HMI tags "BC_HMI_Tags"
   "10 DI_DATA_E131_OK" : Bool = PLC "20_TANKS_IP_DATA".RIO_03.FIRST_TANK.USD_FLOW AT %DB1.DBX0.0, 1 s
   "10 DI_DATA_E131_SHTDN" : Bool = PLC "10 DI_DATA".E131_SHTDN AT %DB1.DBX0.0, 1 s
   "103_Main_Burner_DB_DN_OK(1)" : Bool = PLC "103_Main_Burner_DB".DN_OK AT %DB1.DBX0.0, 1 s
   "10 DI_DATA_FD001_OK" : Bool = PLC "10 DI_DATA".FD001_OK AT %DB1.DBX0.0, 1 s
   "10 DI_DATA_FD001_PWR_OK" : Bool = PLC "10 DI_DATA".FD001_PWR_OK AT %DB1.DBX0.0, 1 s
   "10 DI_DATA_FS115(1)" : Bool = PLC "10 DI_DATA".FS115 AT %DB1.DBW0, 1 s
   "10 DI_DATA_FS123" : Bool = PLC "10 DI_DATA".FS123 AT %DB1.DBX0.0, 1 s
   "10 DI_DATA_FS317" : Bool = PLC "10 DI_DATA".FS317 AT %DB1.DBX0.0, 1 s
   "10 DI_DATA_FS320" : Bool = PLC "10 DI_DATA".FS320 AT %DB1.DBX0.0, 1 s
   "10 DI_DATA_ESD_OK" : Bool = PLC "10 DI_DATA".ESD_OK AT %DB1.DBX0.0, 1 s
   "10 DI_DATA_P301_ENBLD" : Bool = PLC "10 DI_DATA".P301_ENBLD AT %DB1.DBX0.0, 1 s
   "10 DI_DATA_R2_SPR_DI_1_6" : Bool = PLC "10 DI_DATA".R2_SPR_DI_1_6 AT %DB1.DBX0.0, 1 s
   "10 DI_DATA_P301_TRIPPED(1)" : Bool = PLC "10 DI_DATA".P301_TRIPPED AT %DB1.DBX0.0, 1 s
   "10 DI_DATA_P305_ENBLD" : Bool = PLC "10 DI_DATA".P305_ENBLD AT %DB1.DBX0.0, 1 s
   "10 DI_DATA_P305_TRIPPED(1)" : Bool = PLC "10 DI_DATA".P305_TRIPPED AT %DB1.DBX0.0, 1 s
   "10 DI_DATA_PS101" : Bool = PLC "10 DI_DATA".PS101 AT %DB1.DBX0.0, 1 s
   "10 DI_DATA_R2_SPR_DI_0_2" : Bool = PLC "10 DI_DATA".R2_SPR_DI_0_2 AT %DB1.DBX0.0, 1 s
   "10 DI_DATA_R2_SPR_DI_0_3" : Bool = PLC "10 DI_DATA".R2_SPR_DI_0_3 AT %DB1.DBX0.0, 1 s
   "10 DI_DATA_TS403_FAULT" : Bool = PLC "10 DI_DATA".TS403_FAULT AT %DB1.DBX0.0, 1 s
   "10 DI_DATA_X001_PWR_OK" : Bool = PLC "10 DI_DATA".X001_PWR_OK AT %DB1.DBX0.0, 1 s
   "102_Pilot_Burner_DB_FLM_DET" : Bool = PLC "102_Pilot_Burner_DB".FLM_DET AT %DB1.DBX0.0, 100 ms
   "104_Pilot_Purge_DB_DN_OK" : Bool = PLC "104_Pilot_Purge_DB".DN_OK AT %DB1.DBX0.0, 1 s
   "10 DI_DATA_E600_NOK" : Bool = PLC "10 DI_DATA".E600_NOK AT %DB1.DBX0.0, 1 s
   "10 DI_DATA_E600_HIHI" : Bool = PLC "10 DI_DATA".E600_HIHI AT %DB1.DBX0.0, 1 s
   "10 DI_DATA_E600_LOLO" : Bool = PLC "10 DI_DATA".E600_LOLO AT %DB1.DBX0.0, 1 s
   "10 DI_DATA_E600_PWR_OK" : Bool = PLC "10 DI_DATA".E600_PWR_OK AT %DB1.DBX0.0, 1 s
   "10 DI_DATA_E700_PWR_OK" : Bool = PLC "10 DI_DATA".E700_PWR_OK AT %DB1.DBX0.0, 1 s
   "10 DI_DATA_E700_OPACITY" : Bool = PLC "10 DI_DATA".E700_OPACITY AT %DB1.DBX0.0, 1 s
   "10 DI_DATA_TS403_FAULT(1)" : Bool = PLC "10 DI_DATA".TS403_FAULT AT %DB1.DBX0.0, 1 s
   "10 DI_DATA_TS006" : Bool = PLC "10 DI_DATA".TS006 AT %DB1.DBX0.0, 1 s
   "10 DI_DATA_S2_8K1_OK" : Bool = PLC "10 DI_DATA".S2_8K1_OK AT %DB1.DBX0.0, 1 s
   "10 DI_DATA_E131_WRNG" : Bool = PLC "10 DI_DATA".E131_WRNG AT %DB1.DBX0.0, 1 s
   "10 DI_DATA_R2_SPR_DI_3_2" : Bool = PLC "10 DI_DATA".R2_SPR_DI_3_2 AT %DB1.DBX0.0, 1 s
   "10 DI_DATA_R2_SPR_DI_3_7" : Bool = PLC "10 DI_DATA".R2_SPR_DI_3_7 AT %DB1.DBX0.0, 1 s
   "10 DI_DATA_LS001" : Bool = PLC "10 DI_DATA".LS001 AT %DB1.DBX0.0, 1 s
   "10 DI_DATA_P305_TRIPPED" : Bool = PLC "10 DI_DATA".P305_TRIPPED AT %DB1.DBX0.0, 1 s
   "10 DI_DATA_P305_ENBLD(1)" : Bool = PLC "10 DI_DATA".P305_ENBLD AT %DB1.DBX0.0, 1 s
   "84_Setpoints_PIT113_High" : Real = PLC "84_Setpoints".PIT113_High AT %DB1.DBD0, 1 s
   "84_Setpoints_PIT113_HighHigh" : Real = PLC "84_Setpoints".PIT113_HighHigh AT %DB1.DBD0, 1 s
   "84_Setpoints_PIT113_Pilot_Target" : Real = PLC "84_Setpoints".PIT113_Pilot_Target AT %DB1.DBX0.0, 1 s
   "84_Setpoints_PIT204_High(2)" : Real = PLC "84_Setpoints".PIT204_High, 1 s
   "84_Setpoints_PIT204_HighHigh(2)" : Real = PLC "84_Setpoints".PIT204_HighHigh, 1 s
   "84_Setpoints_PIT204_Low(2)" : Real = PLC "84_Setpoints".PIT204_Low, 1 s
   "84_Setpoints_PIT204_LowLow(2)" : Real = PLC "84_Setpoints".PIT204_LowLow, 1 s
   "84_Setpoints_PIT205_High" : Real = PLC "2084_Setpoints"."TX427 Star DO Lo" AT %DB1.DBD0, 1 s
   "84_Setpoints_PIT205_HighHigh" : Real = PLC "84_Setpoints".PIT205_HighHigh AT %DB1.DBD0, 1 s
   "84_Setpoints_PIT205_Low" : Real = PLC "84_Setpoints".PIT205_Low AT %DB1.DBD0, 1 s
   "84_Setpoints_PIT205_LowLow" : Real = PLC "84_Setpoints".PIT205_LowLow AT %DB1.DBD0, 1 s
   "84_Setpoints_PIT205_Target" : Real = PLC "84_Setpoints".PIT205_Target AT %DB1.DBX0.0, 1 s
   "84_Setpoints_PIT113_Low" : Real = PLC "84_Setpoints".PIT113_Low AT %DB1.DBD0, 1 s
   "84_Setpoints_PIT113_LowLow" : Real = PLC "84_Setpoints".PIT113_LowLow AT %DB1.DBD0, 1 s
   "84_Setpoints_TIT202_High" : Real = PLC "84_Setpoints".TIT202_High AT %DB1.DBD0, 1 s
   "84_Setpoints_TIT202_HighHigh" : Real = PLC "84_Setpoints".TIT202_HighHigh AT %DB1.DBD0, 1 s
   "84_Setpoints_TIT202_LowLow" : Real = PLC "84_Setpoints".TIT202_LowLow AT %DB1.DBD0, 1 s
   "84_Setpoints_TIT202_Low" : Real = PLC "84_Setpoints".TIT202_Low AT %DB1.DBD0, 1 s
   "84_Setpoints_TX700_High" : Real = PLC "84_Setpoints".TX700_High AT %DB1.DBD0, 1 s
   "84_Setpoints_TX700_Low" : Real = PLC "84_Setpoints".TX700_Low AT %DB1.DBD0, 1 s
   "84_Setpoints_FD001_LowLow" : Real = PLC "84_Setpoints".FD001_LowLow AT %DB1.DBD0, 1 s
   "84_Setpoints_E600_BWT_High" : Real = PLC "84_Setpoints".E600_BWT_High AT %DB1.DBD0, 1 s
   "84_Setpoints_E600_BWT_Low" : Real = PLC "84_Setpoints".E600_BWT_Low AT %DB1.DBD0, 1 s
   "84_Setpoints_FD001_Low" : Real = PLC "84_Setpoints".FD001_Low AT %DB1.DBD0, 1 s
   "84_Setpoints_AT_O2_1_LowLow" : Real = PLC "84_Setpoints".AT_O2_1_LowLow AT %DB1.DBD0, 1 s
   "84_Setpoints_AT_O2_2_LowLow" : Real = PLC "84_Setpoints".AT_O2_2_LowLow AT %DB1.DBD0, 1 s
   "84_Setpoints_AT_O2_2_Low" : Real = PLC "84_Setpoints".AT_O2_2_Low AT %DB1.DBD0, 1 s
   "80_From_HMI_MAN_DQ_1_7(1)" : Bool = PLC "80_From_HMI".MAN_DQ_1_7 AT %DB1.DBX0.0, 1 s
   "80_From_HMI_MAN_DQ_1_6" : Bool = PLC "80_From_HMI".MAN_DQ_1_6 AT %DB1.DBX0.0, 1 s
   "80_From_HMI_MAN_DQ_1_5(1)" : Bool = PLC "80_From_HMI".MAN_DQ_1_5 AT %DB1.DBX0.0, 1 s
   "80_From_HMI_MAN_DQ_1_4(1)" : Bool = PLC "80_From_HMI".MAN_DQ_1_4 AT %DB1.DBX0.0, 1 s
   "80_From_HMI_MAN_DQ_1_3(1)" : Bool = PLC "80_From_HMI".MAN_DQ_1_3 AT %DB1.DBX0.0, 1 s
   "80_From_HMI_MAN_DQ_1_2(1)" : Bool = PLC "80_From_HMI".MAN_DQ_1_2 AT %DB1.DBX0.0, 1 s
   "80_From_HMI_MAN_DQ_1_1(1)" : Bool = PLC "80_From_HMI".MAN_DQ_1_1 AT %DB1.DBX0.0, 1 s
   "80_From_HMI_MAN_DQ_1_0" : Bool = PLC "80_From_HMI".MAN_DQ_1_0 AT %DB1.DBX0.0, 1 s
   "80_From_HMI_MAN_DQ_0_7" : Bool = PLC "80_From_HMI".MAN_DQ_0_7 AT %DB1.DBX0.0, 1 s
   "80_From_HMI_MAN_DQ_0_6(1)" : Bool = PLC "80_From_HMI".MAN_DQ_0_6 AT %DB1.DBX0.0, 1 s
   "80_From_HMI_MAN_DQ_0_5(1)" : Bool = PLC "80_From_HMI".MAN_DQ_0_5 AT %DB1.DBX0.0, 1 s
   "80_From_HMI_MAN_DQ_0_4(1)" : Bool = PLC "80_From_HMI".MAN_DQ_0_4 AT %DB1.DBX0.0, 1 s
   "80_From_HMI_MAN_DQ_0_3(1)" : Bool = PLC "80_From_HMI".MAN_DQ_0_3 AT %DB1.DBX0.0, 1 s
   "80_From_HMI_MAN_DQ_0_2(1)" : Bool = PLC "80_From_HMI".MAN_DQ_0_2 AT %DB1.DBX0.0, 1 s
   "80_From_HMI_MAN_DQ_0_1(1)" : Bool = PLC "80_From_HMI".MAN_DQ_0_1 AT %DB1.DBX0.0, 1 s
   "80_From_HMI_MAN_DQ_0_0(1)" : Bool = PLC "80_From_HMI".MAN_DQ_0_0 AT %DB1.DBX0.0, 1 s
   "16_AQ_Data_CV111_CNTRL" : Real = PLC "16_AQ_Data".CV111_CNTRL AT %DB1.DBD0, 1 s
   "14_DQ_Data_X001ControlOut" : Bool = PLC "14_DQ_Data".X001ControlOut AT %DB1.DBX0.0, 1 s
   "14_DQ_Data_R2_SPR_DQ_1_6" : Bool = PLC "14_DQ_Data".R2_SPR_DQ_1_6 AT %DB1.DBX0.0, 1 s
   "14_DQ_Data_R2_SPR_DQ_1_4" : Bool = PLC "14_DQ_Data".R2_SPR_DQ_1_4 AT %DB1.DBX0.0, 1 s
   "14_DQ_Data_R2_SPR_DQ_1_5" : Bool = PLC "14_DQ_Data".R2_SPR_DQ_1_5 AT %DB1.DBX0.0, 1 s
   "14_DQ_Data_R2_SPR_DQ_1_3" : Bool = PLC "14_DQ_Data".R2_SPR_DQ_1_3 AT %DB1.DBX0.0, 1 s
   "14_DQ_Data_R2_SPR_DQ_1_2" : Bool = PLC "14_DQ_Data".R2_SPR_DQ_1_2 AT %DB1.DBX0.0, 1 s
   "14_DQ_Data_P305ControlOut" : Bool = PLC "14_DQ_Data".P305ControlOut AT %DB1.DBX0.0, 1 s
   "14_DQ_Data_E131ControlOut" : Bool = PLC "14_DQ_Data".E131ControlOut AT %DB1.DBX0.0, 1 s
   "14_DQ_Data_200CV216ControlOut" : Bool = PLC "14_DQ_Data".200CV216ControlOut AT %DB1.DBX0.0, 1 s
   "14_DQ_Data_200CV215ControlOut" : Bool = PLC "14_DQ_Data".200CV215ControlOut AT %DB1.DBX0.0, 1 s
   "14_DQ_Data_200CV207ControlOut" : Bool = PLC "14_DQ_Data".200CV207ControlOut AT %DB1.DBX0.0, 1 s
   "14_DQ_Data_200CV206ControlOut" : Bool = PLC "14_DQ_Data".200CV206ControlOut AT %DB1.DBX0.0, 1 s
   "14_DQ_Data_200CV127ControlOut" : Bool = PLC "14_DQ_Data".200CV127ControlOut AT %DB1.DBX0.0, 1 s
   "14_DQ_Data_200CV124ControlOut" : Bool = PLC "14_DQ_Data".200CV124ControlOut AT %DB1.DBX0.0, 1 s
   "14_DQ_Data_200CV114ControlOut" : Bool = PLC "14_DQ_Data".200CV114ControlOut AT %DB1.DBX0.0, 1 s
   "12_AI_Data_TIT202In_SCALED" : Real = PLC "12_AI_Data".TIT202In_SCALED AT %DB1.DBX0.0, 1 s
   "12_AI_Data_PIT205In_SCALED" : Real = PLC "12_AI_Data".PIT205In_SCALED AT %DB1.DBX0.0, 1 s
   "12_AI_Data_PIT204In_SCALED" : Real = PLC "12_AI_Data".PIT204In_SCALED AT %DB1.DBX0.0, 1 s
   "12_AI_Data_PIT112In_SCALED" : Real = PLC "12_AI_Data".PIT112In_SCALED AT %DB1.DBX0.0, 1 s
   "12_AI_Data_FD001FlameSignalIn" : Real = PLC "12_AI_Data".FD001FlameSignalIn AT %DB1.DBX0.0, 100 ms
   "12_AI_Data_E700SootContentIn" : Real = PLC "12_AI_Data".E700SootContentIn AT %DB1.DBX0.0, 1 s
   "12_AI_Data_E600O2ContentIn" : Real = PLC "12_AI_Data".E600O2ContentIn AT %DB1.DBX0.0, 100 ms
   "10 DI_DATA_TS403_FAULT(2)" : Bool = PLC "10 DI_DATA".TS403_FAULT AT %DB1.DBX0.0, 1 s
   "10_DI_Data_E139_RUNNING" : Bool = PLC "10_DI_Data".E139_RUNNING AT %DB1.DBX0.0, 1 s
   "10 DI_DATA_TS006(1)" : Bool = PLC "10 DI_DATA".TS006 AT %DB1.DBX0.0, 1 s
   "16_AQ_Data_CV203_CNTRL" : Real = PLC "16_AQ_Data".CV203_CNTRL AT %DB1.DBD0, 1 s
   "16_AQ_Data_R2_SPR_AQ_96" : Real = PLC "16_AQ_Data".R2_SPR_AQ_96 AT %DB1.DBD0, 1 s
   "16_AQ_Data_R2_SPR_AQ_98" : Real = PLC "16_AQ_Data".R2_SPR_AQ_98 AT %DB1.DBD0, 1 s
   "80_From_HMI_MAN_AQ_INC_96" : Bool = PLC "80_From_HMI".MAN_AQ_INC_96 AT %DB1.DBX0.0, 1 s
   "80_From_HMI_MAN_AQ_DEC_96" : Bool = PLC "80_From_HMI".MAN_AQ_DEC_96 AT %DB1.DBX0.0, 1 s
   "80_From_HMI_MAN_AQ_INC_98" : Bool = PLC "80_From_HMI".MAN_AQ_INC_98 AT %DB1.DBX0.0, 1 s
   "80_From_HMI_MAN_AQ_DEC_98" : Bool = PLC "80_From_HMI".MAN_AQ_DEC_98 AT %DB1.DBX0.0, 1 s
   "80_From_HMI_MAN_AQ_INC_100(1)" : Bool = PLC "80_From_HMI".MAN_AQ_INC_100 AT %DB1.DBX0.0, 1 s
   "80_From_HMI_MAN_AQ_DEC_100(1)" : Bool = PLC "80_From_HMI".MAN_AQ_DEC_100 AT %DB1.DBX0.0, 1 s
   "80_From_HMI_MAN_AQ_INC_102" : Bool = PLC "80_From_HMI".MAN_AQ_INC_102 AT %DB1.DBX0.0, 1 s
   "80_From_HMI_MAN_AQ_DEC_102" : Bool = PLC "80_From_HMI".MAN_AQ_DEC_102 AT %DB1.DBX0.0, 1 s
   "10 DI_DATA_FS115" : Bool = PLC "10 DI_DATA".FS115 AT %DB1.DBX0.0, 1 s
   "10 DI_DATA_P301_TRIPPED" : Bool = PLC "10 DI_DATA".P301_TRIPPED AT %DB1.DBX0.0, 1 s
   "84_Setpoints_E600_BWT_HighHigh" : Real = PLC "84_Setpoints".E600_BWT_HighHigh AT %DB1.DBD0, 1 s
   "84_Setpoints_E600_BWT_LowLow" : Real = PLC "84_Setpoints".E600_BWT_LowLow AT %DB1.DBD0, 1 s
   "84_Setpoints_E600_CB_Low" : Real = PLC "84_Setpoints".E600_CB_Low AT %DB1.DBD0, 1 s
   "84_Setpoints_E600_CB_LowLow" : Real = PLC "84_Setpoints".E600_CB_LowLow AT %DB1.DBD0, 1 s
   "84_Setpoints_E600_CB_High" : Real = PLC "84_Setpoints".E600_CB_High AT %DB1.DBD0, 1 s
   "84_Setpoints_E600_CB_HighHigh" : Real = PLC "84_Setpoints".E600_CB_HighHigh AT %DB1.DBD0, 1 s
   "84_Setpoints_FD001_Min" : Real = PLC "84_Setpoints".FD001_Min AT %DB1.DBD0, 1 s
   "84_Setpoints_PIT113_Pilot_Target(1)" : Real = PLC "62_Warning_Data".GCU_WARNING_WORD_01 AT %DB1.DBD0, 1 s
   "84_Setpoints_PIT205_Target(1)" : Real = PLC "84_Setpoints".PIT205_Target AT %DB1.DBD0, 1 s
   "84_Setpoints_E600_CB_Target" : Real = PLC "84_Setpoints".E600_CB_Target AT %DB1.DBD0, 1 s
   "84_Setpoints_E600_BWT_Target" : Real = PLC "84_Setpoints".E600_BWT_Target AT %DB1.DBD0, 1 s
   "86_Times_CV127_OPEN_TIME_#1" : Time = PLC "86_Times".CV127_OPEN_TIME_#1 AT %DB1.DBX0.0, 1 s
   "86_Times_CV127_CLOSED_TIME" : Time = PLC "86_Times".CV127_CLOSED_TIME AT %DB1.DBX0.0, 1 s
   "86_Times_CV127_OPEN_TIME_#2" : Time = PLC "86_Times".CV127_OPEN_TIME_#2 AT %DB1.DBX0.0, 1 s
   "86_Times_CV124_OPEN_TIME" : Time = PLC "86_Times".CV124_OPEN_TIME AT %DB1.DBX0.0, 1 s
   "86_Times_CV124_CLOSE_TIME_PRG" : Time = PLC "86_Times".CV124_CLOSE_TIME_PRG AT %DB1.DBX0.0, 1 s
   "86_Times_CV114_OPEN_TIME" : Time = PLC "86_Times".CV114_OPEN_TIME AT %DB1.DBX0.0, 1 s
   "86_Times_CV206_OPEN_TIME" : Time = PLC "86_Times".CV206_OPEN_TIME AT %DB1.DBX0.0, 1 s
   "86_Times_CV207_OPEN_TIME" : Time = PLC "86_Times".CV207_OPEN_TIME AT %DB1.DBX0.0, 1 s
   "86_Times_CV215_OPEN_TIME" : Time = PLC "86_Times".CV215_OPEN_TIME AT %DB1.DBX0.0, 1 s
   "86_Times_CV215_CLOSE_TIME_PRG" : Time = PLC "86_Times".CV215_CLOSE_TIME_PRG AT %DB1.DBX0.0, 1 s
   "86_Times_CV216_OPEN_TIME" : Time = PLC "86_Times".CV216_OPEN_TIME AT %DB1.DBX0.0, 1 s
   "86_Times_CV216_CLOSE_TIME_PRG" : Time = PLC "86_Times".CV216_CLOSE_TIME_PRG AT %DB1.DBX0.0, 1 s
   "86_Times_CV216_OPEN_TIME_PRG" : Time = PLC "86_Times".CV216_OPEN_TIME_PRG AT %DB1.DBX0.0, 1 s
   "86_Times_CV206_CLOSE_TIME" : Time = PLC "86_Times".CV206_CLOSE_TIME AT %DB1.DBX0.0, 1 s
   "86_Times_CV207_CLOSE_TIME" : Time = PLC "86_Times".CV207_CLOSE_TIME AT %DB1.DBX0.0, 1 s
   "86_Times_CV114_CLOSE_TIME" : Time = PLC "86_Times".CV114_CLOSE_TIME AT %DB1.DBD0, 1 s
   "86_Times_CV215_CLOSE_TIME" : Time = PLC "86_Times".CV215_CLOSE_TIME AT %DB1.DBD0, 1 s
   "86_Times_CV216_CLOSE_TIME" : Time = PLC "86_Times".CV216_CLOSE_TIME AT %DB1.DBD0, 1 s
   "86_Times_CV124_CLOSE_TIME" : Time = PLC "86_Times".CV124_CLOSE_TIME AT %DB1.DBD0, 1 s
   "86_Times_X001_MAX_RUN_TIME" : Time = PLC "86_Times".X001_MAX_RUN_TIME AT %DB1.DBD0, 1 s
   "86_Times_X001_RUN_CNF_TIME" : Time = PLC "86_Times".X001_RUN_CNF_TIME AT %DB1.DBD0, 1 s
   "86_Times_FD_DET_DELAY" : Time = PLC "86_Times".FD_DET_DELAY AT %DB1.DBD0, 1 s
   "86_Times_FD_VRFCTN_TIME" : Time = PLC "86_Times".FD_VRFCTN_TIME AT %DB1.DBD0, 1 s
   "86_Times_FDU_DET_TIME" : Time = PLC "86_Times".FDU_DET_TIME AT %DB1.DBD0, 1 s
   "86_Times_MAX_IGNTN_SEQ_TIME" : Time = PLC "86_Times".MAX_IGNTN_SEQ_TIME AT %DB1.DBD0, 1 s
   "86_Times_MAX_MAIN_BURN_SEQ_TIME" : Time = PLC "86_Times".MAX_MAIN_BURN_SEQ_TIME AT %DB1.DBD0, 1 s
   "86_Times_MAX_PILOT_PURGE_SEQ_TIME" : Time = PLC "86_Times".MAX_PILOT_PURGE_SEQ_TIME AT %DB1.DBD0, 1 s
   "86_Times_O2_CHECK_TIME" : Time = PLC "86_Times".O2_CHECK_TIME AT %DB1.DBD0, 1 s
   "86_Times_STEP_MAX_TIME_STP_001(1)" : Time = PLC "86_Times".STEP_MAX_TIME_STP_001 AT %DB1.DBW0, 1 s
   "86_Times_STEP_MAX_TIME_STP_005(1)" : Time = PLC "86_Times".STEP_MAX_TIME_STP_005 AT %DB1.DBW0, 1 s
   "86_Times_STEP_MAX_TIME_STP_010(1)" : Time = PLC "86_Times".STEP_MAX_TIME_STP_010 AT %DB1.DBW0, 1 s
   "86_Times_STEP_MAX_TIME_STP_020(1)" : Time = PLC "86_Times".STEP_MAX_TIME_STP_020 AT %DB1.DBW0, 1 s
   "86_Times_STEP_MAX_TIME_STP_030(1)" : Time = PLC "86_Times".STEP_MAX_TIME_STP_030 AT %DB1.DBW0, 1 s
   "86_Times_STEP_MAX_TIME_STP_040(1)" : Time = PLC "86_Times".STEP_MAX_TIME_STP_040 AT %DB1.DBW0, 1 s
   "86_Times_STEP_MAX_TIME_STP_050(1)" : Time = PLC "86_Times".STEP_MAX_TIME_STP_050 AT %DB1.DBW0, 1 s
   "86_Times_STEP_MAX_TIME_STP_060(1)" : Time = PLC "86_Times".STEP_MAX_TIME_STP_060 AT %DB1.DBW0, 1 s
   "86_Times_STEP_MAX_TIME_STP_070(1)" : Time = PLC "86_Times".STEP_MAX_TIME_STP_070 AT %DB1.DBW0, 1 s
   "86_Times_STEP_MAX_TIME_STP_080(1)" : Time = PLC "86_Times".STEP_MAX_TIME_STP_080 AT %DB1.DBW0, 1 s
   "86_Times_STEP_MAX_TIME_STP_090(1)" : Time = PLC "86_Times".STEP_MAX_TIME_STP_090 AT %DB1.DBW0, 1 s
   "86_Times_STEP_MAX_TIME_STP_100(1)" : Time = PLC "86_Times".STEP_MAX_TIME_STP_100 AT %DB1.DBW0, 1 s
   "86_Times_STEP_MAX_TIME_STP_110(1)" : Time = PLC "86_Times".STEP_MAX_TIME_STP_110 AT %DB1.DBW0, 1 s
   "86_Times_STEP_MAX_TIME_STP_120(1)" : Time = PLC "86_Times".STEP_MAX_TIME_STP_120 AT %DB1.DBW0, 1 s
   "86_Times_STEP_MAX_TIME_STP_130(1)" : Time = PLC "86_Times".STEP_MAX_TIME_STP_130 AT %DB1.DBW0, 1 s
   "86_Times_STEP_MAX_TIME_STP_140(1)" : Time = PLC "86_Times".STEP_MAX_TIME_STP_140 AT %DB1.DBW0, 1 s
   "86_Times_STEP_MAX_TIME_STP_150(1)" : Time = PLC "86_Times".STEP_MAX_TIME_STP_150 AT %DB1.DBW0, 1 s
   "86_Times_STEP_MAX_TIME_STP_160(1)" : Time = PLC "86_Times".STEP_MAX_TIME_STP_160 AT %DB1.DBW0, 1 s
   "86_Times_STEP_MAX_TIME_STP_170(1)" : Time = PLC "86_Times".STEP_MAX_TIME_STP_170 AT %DB1.DBW0, 1 s
   "86_Times_STEP_MAX_TIME_STP_180(1)" : Time = PLC "86_Times".STEP_MAX_TIME_STP_180 AT %DB1.DBW0, 1 s
   "86_Times_STEP_MAX_TIME_STP_190(1)" : Time = PLC "86_Times".STEP_MAX_TIME_STP_190 AT %DB1.DBW0, 1 s
   "86_Times_STEP_MAX_TIME_STP_200(1)" : Time = PLC "86_Times".STEP_MAX_TIME_STP_200 AT %DB1.DBW0, 1 s
   "86_Times_STEP_MAX_TIME_STP_210(1)" : Time = PLC "86_Times".STEP_MAX_TIME_STP_210 AT %DB1.DBW0, 1 s
   "86_Times_STEP_MAX_TIME_STP_220(1)" : Time = PLC "86_Times".STEP_MAX_TIME_STP_220 AT %DB1.DBW0, 1 s
   "86_Times_STEP_MAX_TIME_STP_230(1)" : Time = PLC "86_Times".STEP_MAX_TIME_STP_230 AT %DB1.DBW0, 1 s
   "86_Times_STEP_MAX_TIME_STP_240(1)" : Time = PLC "86_Times".STEP_MAX_TIME_STP_240 AT %DB1.DBW0, 1 s
   "86_Times_STEP_MAX_TIME_STP_250(1)" : Time = PLC "86_Times".STEP_MAX_TIME_STP_250 AT %DB1.DBW0, 1 s
   "86_Times_STEP_MAX_TIME_STP_260(1)" : Time = PLC "86_Times".STEP_MAX_TIME_STP_260 AT %DB1.DBW0, 1 s
   "86_Times_STEP_MAX_TIME_STP_270(1)" : Time = PLC "86_Times".STEP_MAX_TIME_STP_270 AT %DB1.DBW0, 1 s
   "86_Times_STEP_MAX_TIME_STP_280(1)" : Time = PLC "86_Times".STEP_MAX_TIME_STP_280 AT %DB1.DBW0, 1 s
   "86_Times_STEP_MAX_TIME_STP_290(1)" : Time = PLC "86_Times".STEP_MAX_TIME_STP_290 AT %DB1.DBW0, 1 s
   "86_Times_STEP_MAX_TIME_STP_300(1)" : Time = PLC "86_Times".STEP_MAX_TIME_STP_300 AT %DB1.DBW0, 1 s
   "86_Times_STEP_MAX_TIME_STP_310(1)" : Time = PLC "86_Times".STEP_MAX_TIME_STP_310 AT %DB1.DBW0, 1 s
   "86_Times_STEP_MAX_TIME_STP_320(1)" : Time = PLC "86_Times".STEP_MAX_TIME_STP_320 AT %DB1.DBW0, 1 s
   "86_Times_STEP_MAX_TIME_STP_330(1)" : Time = PLC "86_Times".STEP_MAX_TIME_STP_330 AT %DB1.DBW0, 1 s
   "86_Times_STEP_MAX_TIME_STP_340(1)" : Time = PLC "86_Times".STEP_MAX_TIME_STP_340 AT %DB1.DBW0, 1 s
   "86_Times_STEP_MAX_TIME_STP_350(1)" : Time = PLC Alarms_Acknowledge.IGG_ALARM_ACKNLG_2 AT %DB1.DBW0, 1 s
   "86_Times_STEP_MAX_TIME_STP_360(1)" : Time = PLC "86_Times".STEP_MAX_TIME_STP_360 AT %DB1.DBW0, 1 s
   "86_Times_STEP_MAX_TIME_STP_370(1)" : Time = PLC "86_Times".STEP_MAX_TIME_STP_370 AT %DB1.DBW0, 1 s
   "86_Times_STEP_MAX_TIME_STP_380(1)" : Time = PLC "86_Times".STEP_MAX_TIME_STP_380 AT %DB1.DBW0, 1 s
   "86_Times_STEP_MAX_TIME_STP_390(1)" : Time = PLC "86_Times".STEP_MAX_TIME_STP_390 AT %DB1.DBW0, 1 s
   "86_Times_STEP_MAX_TIME_STP_400(1)" : Time = PLC "86_Times".STEP_MAX_TIME_STP_400 AT %DB1.DBW0, 1 s
   "86_Times_STEP_MAX_TIME_STP_410(1)" : Time = PLC "86_Times".STEP_MAX_TIME_STP_410 AT %DB1.DBW0, 1 s
   "86_Times_STEP_MAX_TIME_STP_420(1)" : Time = PLC "86_Times".STEP_MAX_TIME_STP_420 AT %DB1.DBW0, 1 s
   "86_Times_STEP_MAX_TIME_STP_430(1)" : Time = PLC "86_Times".STEP_MAX_TIME_STP_430 AT %DB1.DBW0, 1 s
   "86_Times_STEP_MAX_TIME_STP_440(1)" : Time = PLC "86_Times".STEP_MAX_TIME_STP_440 AT %DB1.DBW0, 1 s
   "86_Times_STEP_MAX_TIME_STP_450(1)" : Time = PLC "86_Times".STEP_MAX_TIME_STP_450 AT %DB1.DBW0, 1 s
   "86_Times_STEP_MAX_TIME_STP_460(1)" : Time = PLC "86_Times".STEP_MAX_TIME_STP_460 AT %DB1.DBW0, 1 s
   "86_Times_STEP_MAX_TIME_STP_470(1)" : Time = PLC "86_Times".STEP_MAX_TIME_STP_470 AT %DB1.DBW0, 1 s
   "86_Times_STEP_MAX_TIME_STP_480(1)" : Time = PLC "86_Times".STEP_MAX_TIME_STP_480 AT %DB1.DBW0, 1 s
   "86_Times_STEP_MAX_TIME_STP_490(1)" : Time = PLC "86_Times".STEP_MAX_TIME_STP_490 AT %DB1.DBW0, 1 s
   "86_Times_STEP_MAX_TIME_STP_500(1)" : Time = PLC "86_Times".STEP_MAX_TIME_STP_500 AT %DB1.DBW0, 1 s
   "86_Times_STEP_MAX_TIME_STP_510(1)" : Time = PLC "86_Times".STEP_MAX_TIME_STP_510 AT %DB1.DBW0, 1 s
   "86_Times_STEP_MAX_TIME_STP_520(1)" : Time = PLC "86_Times".STEP_MAX_TIME_STP_520 AT %DB1.DBW0, 1 s
   "86_Times_STEP_MAX_TIME_STP_530(1)" : Time = PLC "86_Times".STEP_MAX_TIME_STP_530 AT %DB1.DBW0, 1 s
   "86_Times_STEP_MAX_TIME_STP_540(1)" : Time = PLC "86_Times".STEP_MAX_TIME_STP_540 AT %DB1.DBW0, 1 s
   "86_Times_STEP_MAX_TIME_STP_550(1)" : Time = PLC "86_Times".STEP_MAX_TIME_STP_550 AT %DB1.DBW0, 1 s
   "86_Times_STEP_MAX_TIME_STP_560(1)" : Time = PLC "86_Times".STEP_MAX_TIME_STP_560 AT %DB1.DBW0, 1 s
   "86_Times_STEP_MAX_TIME_STP_570(1)" : Time = PLC "10_DI_DATA".R3_SPR_DI_136_0 AT %DB1.DBW0, 1 s

HMI tags "IGG_HMI_Tags"
   "10_DI_Data_CV311_OPN" : Bool = PLC "10_DI_Data".CV311_OPN AT %DB1.DBW0, 1 s
   "10_DI_Data_CV311_CLSD" : Bool = PLC "82_To_HMI"."I&A Compressor Service Due" AT %DB1.DBW0, 1 s
   "80_From_HMI_RUN_IGG" : Bool = PLC "80_From_HMI".RUN_IGG AT %DB1.DBX0.0, 1 s
   "82_To_HMI_CA Blower Animation" : Int = PLC "82_To_HMI"."CA Blower Animation" AT %DB1.DBX0.0, 100 ms
   "10_DI_Data_E500B_ENBLD" : Bool = PLC "10_DI_Data".E500B_ENBLD AT %DB1.DBX0.0, 1 s
   "10_DI_Data_E500A_ENBLD" : Bool = PLC "10_DI_Data".E500A_ENBLD AT %DB1.DBX0.0, 1 s
   "80_From_HMI_RUN_IGG(1)" : Bool = PLC "80_From_HMI".RUN_IGG AT %DB1.DBX0.0, 1 s
   "14_DQ_Data_E500A_CNTRL" : Bool = PLC "14_DQ_Data".E500A_CNTRL AT %DB1.DBX0.0, 1 s
   "14_DQ_Data_E500B_CNTRL" : Bool = PLC "14_DQ_Data".E500B_CNTRL AT %DB1.DBX0.0, 1 s
   "82_To_HMI_Run Time A" : LTime = PLC "82_To_HMI"."Run Time A" AT %DB1.DBD0, 1 s
   "82_To_HMI_Run Time B" : LTime = PLC "82_To_HMI"."Run Time B" AT %DB1.DBD0, 1 s
   "80_From_HMI_SW_DTY_PMP_E500" : Bool = PLC "80_From_HMI".SW_DTY_PMP_E500 AT %DB1.DBW0, 1 s
   "12_AI_Data_PIT316_SCALED" : Real = PLC "12_AI_Data".PIT316_SCALED AT %DB1.DBX0.0, 1 s
   "12_AI_Data_TIT319_SCALED" : Real = PLC "12_AI_Data".TIT319_SCALED AT %DB1.DBX0.0, 1 s
   "12_AI_Data_TIT360_SCALED" : Real = PLC "12_AI_Data".TIT360_SCALED AT %DB1.DBX0.0, 1 s
   "12_AI_Data_PIT102_SCALED(1)" : Real = PLC "12_AI_Data".PIT102_SCALED AT %DB1.DBX0.0, 1 s
   "12_AI_Data_CV403_SCALED(1)" : Real = PLC "12_AI_Data".CV403_SCALED AT %DB1.DBX0.0, 1 s
   "12_AI_Data_E139_RPM_SCALED" : Real = PLC "12_AI_Data".E139_RPM_SCALED AT %DB1.DBX0.0, 1 s
   "12_AI_Data_E139_AMPS_SCALED" : Real = PLC "12_AI_Data".E139_AMPS_SCALED AT %DB1.DBX0.0, 1 s
   "12_AI_Data_PIT402_SCALED" : Real = PLC "12_AI_Data".PIT402_SCALED AT %DB1.DBX0.0, 1 s
   "10_DI_Data_E500B_TRIPPED" : Bool = PLC "10_DI_Data".E500B_TRIPPED AT %DB1.DBX0.0, 1 s
   "10_DI_Data_IGG_ESTOP_OK" : Bool = PLC "10_DI_Data".IGG_ESTOP_OK AT %DB1.DBX0.0, 1 s
   "10_DI_Data_E500A_TRIPPED" : Bool = PLC "10_DI_Data".E500A_TRIPPED AT %DB1.DBX0.0, 1 s
   "10_DI_Data_E500B_TRIPPED(1)" : Bool = PLC "10_DI_Data".E500B_TRIPPED AT %DB1.DBX0.0, 1 s
   "10_DI_Data_E500A_ENBLD(1)" : Bool = PLC "10_DI_Data".E500A_ENBLD AT %DB1.DBX0.0, 1 s
   "10_DI_Data_E500B_ENBLD(1)" : Bool = PLC "10_DI_Data".E500B_ENBLD AT %DB1.DBX0.0, 1 s
   "10_DI_Data_CV401_OPN" : Bool = PLC "10_DI_Data".CV401_OPN AT %DB1.DBX0.0, 1 s
   "10_DI_Data_CV401_CLSD" : Bool = PLC "10_DI_Data".CV401_CLSD AT %DB1.DBX0.0, 1 s
   "10_DI_Data_CV321_OPN" : Bool = PLC "10_DI_Data".CV321_OPN AT %DB1.DBX0.0, 1 s
   "10_DI_Data_CV321_CLSD" : Bool = PLC "10_DI_Data".CV321_CLSD AT %DB1.DBX0.0, 1 s
   "10_DI_Data_CV322_OPN" : Bool = PLC "10_DI_Data".CV322_OPN AT %DB1.DBX0.0, 1 s
   "10_DI_Data_CV322_CLSD" : Bool = PLC "10_DI_Data".CV322_CLSD AT %DB1.DBX0.0, 1 s
   "10_DI_Data_BC_PLC_PWR_OK" : Bool = PLC "10_DI_Data".BC_PLC_PWR_OK AT %DB1.DBX0.0, 1 s
   "10_DI_Data_IGG_VNT_PWR_OK" : Bool = PLC "10_DI_Data".IGG_VNT_PWR_OK AT %DB1.DBX0.0, 1 s
   "10_DI_Data_MCC_VNT_PWR_OK" : Bool = PLC "10_DI_Data".MCC_VNT_PWR_OK AT %DB1.DBX0.0, 1 s
   "10_DI_Data_7T1_PWR_OK" : Bool = PLC "10_DI_Data".7T1_PWR_OK AT %DB1.DBX0.0, 1 s
   "10_DI_Data_7T2_PWR_OK" : Bool = PLC "10_DI_Data".7T2_PWR_OK AT %DB1.DBX0.0, 1 s
   "10_DI_Data_7T3_PWR_OK" : Bool = PLC "10_DI_Data".7T3_PWR_OK AT %DB1.DBX0.0, 1 s
   "10_DI_Data_MAINTD_24VDC_PWR_OK" : Bool = PLC "10_DI_Data".MAINTD_24VDC_PWR_OK AT %DB1.DBX0.0, 1 s
   "10_DI_Data_SFTY_SYS_IL" : Bool = PLC "10_DI_Data".SFTY_SYS_IL AT %DB1.DBX0.0, 1 s
   "14_DQ_Data_CV311_312_CNTRL" : Bool = PLC "14_DQ_Data".CV311_312_CNTRL AT %DB1.DBX0.0, 1 s
   "14_DQ_Data_CV321_322_CNTRL" : Bool = PLC "14_DQ_Data".CV321_322_CNTRL AT %DB1.DBX0.0, 1 s
   "14_DQ_Data_CV401_CNTRL" : Bool = PLC "14_DQ_Data".CV401_CNTRL AT %DB1.DBX0.0, 1 s
   "51_SLAVE_STATUS_P301_ENBLD" : Bool = PLC "51_SLAVE_STATUS".P301_ENBLD AT %DB51.DBX14.3, 1 s
   "14_DQ_Data_24K2" : Bool = PLC "14_DQ_Data".24K2 AT %DB1.DBX0.0, 1 s
   "14_DQ_Data_24K3" : Bool = PLC "14_DQ_Data".24K3 AT %DB1.DBX0.0, 1 s
   "14_DQ_Data_24K4" : Bool = PLC "14_DQ_Data".24K4 AT %DB1.DBX0.0, 1 s
   "14_DQ_Data_24PF1" : Bool = PLC "14_DQ_Data".24PF1 AT %DB1.DBX0.0, 1 s
   "14_DQ_Data_24K3(2)" : Bool = PLC "14_DQ_Data".24K3 AT %DB1.DBX0.0, 1 s
   "14_DQ_Data_24PF3" : Bool = PLC "14_DQ_Data".24PF3 AT %DB1.DBX0.0, 1 s
   "14_DQ_Data_24PF4" : Bool = PLC "14_DQ_Data".24PF4 AT %DB1.DBX0.0, 100 ms
   "12_AI_Data_PIT102_SCALED" : Real = PLC "12_AI_Data".PIT102_SCALED AT %DB1.DBX0.0, 1 s
   "12_AI_Data_TIT401_SCALED" : Real = PLC "12_AI_Data".TIT401_SCALED AT %DB1.DBX0.0, 1 s
   "12_AI_Data_TIT315_SCALED" : Real = PLC "12_AI_Data".TIT315_SCALED AT %DB1.DBX0.0, 1 s
   "80_From_HMI_Request_Manual(1)" : Bool = PLC "80_From_HMI".Request_Manual AT %DB1.DBX0.0, 1 s
   "12_AI_Data_CV403_SCALED" : Real = PLC "12_AI_Data".CV403_SCALED AT %DB1.DBX0.0, 1 s
   "16_AQ_Data_CV403_CNTRL" : Real = PLC "16_AQ_Data".CV403_CNTRL AT %DB1.DBX0.0, 1 s
   "AlwaysTRUE" : Bool = PLC AlwaysTRUE AT %M1.2, 1 s
   "12_AI_Data_PIT359_SCALED" : Real = PLC "12_AI_Data".PIT359_SCALED AT %DB1.DBX0.0, 1 s
   "68_Sys_Status_Data_CSW_IL_PRES_IN_RNG" : Bool = PLC "68_Sys_Status_Data".CSW_IL_PRES_IN_RNG AT %DB1.DBX0.0, 1 s